// TIA Portal project "DHARMA_1500" (V15) (continued)
VAR_GLOBAL   // PLC tag table "VAT_DeSelectModule"
   "HM_DP_Bus_MK01_Melden" AT %M30.0 : Bool;
   "HM_DP_Bus_MK01_speichern" AT %M30.1 : Bool;
   "HM_DP_Bus_MK01_aktiv" AT %M30.2 : Bool;
   "HM_DP_Bus_MK02_Melden" AT %M30.3 : Bool;
   "HM_DP_Bus_MK02_speichern" AT %M30.4 : Bool;
   "HM_DP_Bus_MK02_aktiv" AT %M30.5 : Bool;
   "HM_DP_Bus_MK03_Melden" AT %M30.6 : Bool;
   "HM_DP_Bus_MK03_speichern" AT %M30.7 : Bool;
   "HM_DP_Bus_MK03_aktiv" AT %M31.0 : Bool;
   "HM_DP_Bus_MK04_Melden" AT %M31.1 : Bool;
   "HM_DP_Bus_MK04_speichern" AT %M31.2 : Bool;
   "HM_DP_Bus_MK04_aktiv" AT %M31.3 : Bool;
   "HM_DP_Bus_MK05_Melden" AT %M31.4 : Bool;
   "HM_DP_Bus_MK05_speichern" AT %M31.5 : Bool;
   "HM_DP_Bus_MK05_aktiv" AT %M31.6 : Bool;
   "HM_DP_Bus_MK06_Melden" AT %M31.7 : Bool;
   "HM_DP_Bus_MK06_speichern" AT %M32.0 : Bool;
   "HM_DP_Bus_MK06_aktiv" AT %M32.1 : Bool;
   "HM_DP_Bus_MK07_Melden" AT %M32.2 : Bool;
   "HM_DP_Bus_MK07_speichern" AT %M32.3 : Bool;
   "HM_DP_Bus_MK07_aktiv" AT %M32.4 : Bool;
   "HM_DP_Bus_MK08_Melden" AT %M32.5 : Bool;
   "HM_DP_Bus_MK08_speichern" AT %M32.6 : Bool;
   "HM_DP_Bus_MK08_aktiv" AT %M32.7 : Bool;
   "HM_DP_Bus_MK09_Melden" AT %M33.0 : Bool;
   "HM_DP_Bus_MK09_speichern" AT %M33.1 : Bool;
   "HM_DP_Bus_MK09_aktiv" AT %M33.2 : Bool;
   "HM_DP_Bus_MK10_Melden" AT %M33.3 : Bool;
   "HM_DP_Bus_MK10_speichern" AT %M33.4 : Bool;
   "HM_DP_Bus_MK10_aktiv" AT %M33.5 : Bool;
   "HM_DP_Bus_MK11_Melden" AT %M33.6 : Bool;
   "HM_DP_Bus_MK11_speichern" AT %M33.7 : Bool;
   "HM_DP_Bus_MK11_aktiv" AT %M34.0 : Bool;
   "HM_DP_Bus_MK12_Melden" AT %M34.1 : Bool;
   "HM_DP_Bus_MK12_speichern" AT %M34.2 : Bool;
   "HM_DP_Bus_MK12_aktiv" AT %M34.3 : Bool;
   "HM_DP_Bus_MK13_Melden" AT %M34.4 : Bool;
   "HM_DP_Bus_MK13_speichern" AT %M34.5 : Bool;
   "HM_DP_Bus_MK13_aktiv" AT %M34.6 : Bool;
   "HM_DP_Bus_MK14_Melden" AT %M34.7 : Bool;
   "HM_DP_Bus_MK14_speichern" AT %M35.0 : Bool;
   "HM_DP_Bus_MK14_aktiv" AT %M35.1 : Bool;
   "HM_DP_Bus_MK15_Melden" AT %M35.2 : Bool;
   "HM_DP_Bus_MK15_speichern" AT %M35.3 : Bool;
   "HM_DP_Bus_MK15_aktiv" AT %M35.4 : Bool;
   "HM_DP_An_Abmelden_Busy" AT %M29.7 : Bool;
END_VAR

VAR_GLOBAL   // PLC tag table "Robots"
   "FHM_PU_cycle_running" AT %M850.0 : Bool;
   "Flag_PU_cycle_running" AT %M850.1 : Bool;
END_VAR

VAR_GLOBAL   // PLC tag table "VAT_VB_Skripte"
   "new_shift" AT %M4.0 : Bool;
   "flag_delay_check_path" AT %M7.1 : Bool;
   "Flag_Network" AT %M1.7 : Bool;
END_VAR

VAR_GLOBAL   // PLC tag table "Shot_protocol"
   "M_ShotActive" AT %M1002.3 : Bool;
   "TotalFlowShotC01" AT %MD950 : Real;
   "TotalFlowShotC02" AT %MD954 : Real;
   "TotalFlowShotC03" AT %MD958 : Real;
   "TotalFlowShotC04" AT %MD962 : Real;
   "TotalFlowShotC05" AT %MD966 : DInt;
   "TotalFlowShotC06" AT %MD970 : DInt;
   "TotalFlowShotC07" AT %MD974 : DInt;
   "TotalFlowShotC08" AT %MD978 : DInt;
   "TotalFlowShotC09" AT %MD982 : DInt;
   "TotalFlowShotC10" AT %MD986 : DInt;
   "TotalFlowShotC11" AT %MD990 : DInt;
   "TotalFlowShotC12" AT %MD994 : DInt;
   "CompAtShot" AT %MW942 : Word;
   "AmountFlowValuesMa1C1" AT %MD800 : Real;
   "AmountFlowValuesMa1C2" AT %MD804 : Real;
   "AmountFlowValuesMa1C3" AT %MD808 : Real;
   "AmountFlowValuesMa1C4" AT %MD812 : Real;
   "FHF_ShotreleaseM1" AT %M940.2 : Bool;
   "M1C01active" AT %M932.0 : Bool;
   "M1C02active" AT %M932.1 : Bool;
   "M1C03active" AT %M932.2 : Bool;
   "M1C04active" AT %M932.3 : Bool;
   "HF_FP_ShotRuns" AT %M941.0 : Bool;
   "HF_FP_ShotStoppedM1" AT %M940.4 : Bool;
   "BufferShotResultM1" AT %M920.0 : Bool;
   "FHM_ShotRunsMH1" AT %M402.0 : Bool;
   "FP_BufferShotResultM1" AT %M919.0 : Bool;
   "M1C05active" AT %M932.4 : Bool;
   "M1C06active" AT %M932.5 : Bool;
   "M1C07active" AT %M932.6 : Bool;
   "M1C08active" AT %M932.7 : Bool;
   "M1C09active" AT %M933.0 : Bool;
   "M1C10active" AT %M933.1 : Bool;
   "M1C11active" AT %M933.2 : Bool;
   "M1C12active" AT %M933.3 : Bool;
   "AmountFlowValuesMa1C5" AT %MD816 : Real;
   "AmountFlowValuesMa1C6" AT %MD820 : Real;
   "AmountFlowValuesMa1C7" AT %MD824 : Real;
   "AmountFlowValuesMa1C8" AT %MD828 : Real;
   "AmountFlowValuesMa1C9" AT %MD832 : Real;
   "AmountFlowValuesMa1C10" AT %MD836 : Real;
   "AmountFlowValuesMa1C11" AT %MD840 : Real;
   "AmountFlowValuesMa1C12" AT %MD844 : Real;
END_VAR

VAR_GLOBAL   // PLC tag table "All_other"
   "TT_Quitt_Door_1" AT %I1102.1 : Bool;
   "TT_H_Empty" AT %Q104.5 : Bool;
   "TT_H_WithoutFoam" AT %Q104.6 : Bool;
   "K_TraceHeatingM1C4" AT %Q16.6 : Bool;
   "Flag_Req_read_DPBus_01" AT %M9.0 : Bool;
   "Flag_Req_read_DP1_Busy" AT %M9.1 : Bool;
   "Flag_Req_read_IO_Busy" AT %M9.2 : Bool;
   "HF_FLT_QPB_C1" AT %M120.1 : Bool;
   "HF_FLT_QPB_C2" AT %M120.2 : Bool;
   "HF_FLT_QPB_C3" AT %M120.3 : Bool;
   "HF_FLT_QPB_C4" AT %M120.4 : Bool;
   "F_CycleRunningMH01" AT %M390.0 : Bool;
   "F_CycleRunningMH02" AT %M390.1 : Bool;
   "F_CycleRunningMH03" AT %M390.2 : Bool;
   "F_CycleRunningMH04" AT %M390.3 : Bool;
   "F_CycleRunningMH05" AT %M390.4 : Bool;
   "F_CycleRunningMH06" AT %M390.5 : Bool;
   "F_CycleRunningMH07" AT %M390.6 : Bool;
   "F_CycleRunningMH08" AT %M390.7 : Bool;
   "StopShotCorrMH01" AT %M309.4 : Bool;
   "StopShotCorrMH02" AT %M309.5 : Bool;
   "StopShotCorrMH03" AT %M309.6 : Bool;
   "StopShotCorrMH04" AT %M309.7 : Bool;
   "ShotFinishedModul_MH01" AT %M122.1 : Bool;
   "ShotFinishedModul_MH02" AT %M122.2 : Bool;
   "ShotFinishedModul_MH03" AT %M122.3 : Bool;
   "ShotFinishedModul_MH04" AT %M122.4 : Bool;
   "ShotFinishedModul_MH05" AT %M122.5 : Bool;
   "ShotFinishedModul_MH06" AT %M122.6 : Bool;
   "ShotFinishedModul_MH07" AT %M122.7 : Bool;
   "ShotFinishedModul_MH08" AT %M123.0 : Bool;
   "ShotFinishedModul_MH09" AT %M123.1 : Bool;
   "ShotFinishedModul_MH10" AT %M123.2 : Bool;
   "ShotFinishedModul_MH11" AT %M123.3 : Bool;
   "ShotFinishedModul_MH12" AT %M123.4 : Bool;
   "ShotFinishedModul_MH13" AT %M123.5 : Bool;
   "ShotFinishedModul_MH14" AT %M123.6 : Bool;
   "ShotFinishedModul_MH15" AT %M123.7 : Bool;
   "ShotFinishedModul_MH16" AT %M124.0 : Bool;
   "EnableFinishShot_MH01" AT %M106.0 : Bool;
   "EnableFinishShot_MH02" AT %M106.1 : Bool;
   "EnableFinishShot_MH03" AT %M106.2 : Bool;
   "EnableFinishShot_MH04" AT %M106.3 : Bool;
   "EnableFinishShot_MH05" AT %M106.4 : Bool;
   "EnableFinishShot_MH06" AT %M106.5 : Bool;
   "EnableFinishShot_MH07" AT %M106.6 : Bool;
   "EnableFinishShot_MH08" AT %M106.7 : Bool;
   "ShotNoNextMa1" AT %MW556 : Int;
   "ShotNoNextMa2" AT %MW558 : Int;
   "ShotNoNextMa3" AT %MW560 : Int;
   "ShotNoNextMa4" AT %MW562 : Int;
   "StopShotCorrMH08" AT %M319.7 : Bool;
   "StopShotCorrMH07" AT %M319.6 : Bool;
   "StopShotCorrMH06" AT %M319.5 : Bool;
   "StopShotCorrMH05" AT %M319.4 : Bool;
   "CalcShotValuesMa1" AT %M135.0 : Bool;
   "ShotStoppedM1" AT %M135.1 : Bool;
   "M1200_ActivateAdrProCan" AT %M120.0 : Bool;
   "NoShotActiveM1" AT %M158.0 : Bool;
   "F_CycleRunningMH09" AT %M391.0 : Bool;
   "F_CycleRunningMH10" AT %M391.1 : Bool;
   "F_CycleRunningMH11" AT %M391.2 : Bool;
   "F_CycleRunningMH12" AT %M391.3 : Bool;
   "F_CycleRunningMH13" AT %M391.4 : Bool;
   "F_CycleRunningMH14" AT %M391.5 : Bool;
   "F_CycleRunningMH15" AT %M391.6 : Bool;
   "F_CycleRunningMH16" AT %M391.7 : Bool;
   "StopShotCorrMH10" AT %M320.1 : Bool;
   "StopShotCorrMH09" AT %M320.0 : Bool;
   "Start_Controler1_HP_K1" AT %M180.5 : Bool;
   "Start_Controler2_HP_K1" AT %M180.4 : Bool;
   "Start_Controler1_HP_K2" AT %M181.5 : Bool;
   "Start_Controler2_HP_K2" AT %M181.4 : Bool;
   "Start_Controler2_LP_K1" AT %M182.4 : Bool;
   "Start_Controler1_LP_K1" AT %M182.5 : Bool;
   "Start_Controler2_LP_K2" AT %M183.4 : Bool;
   "Start_Controler1_LP_K2" AT %M183.5 : Bool;
   "Flag_ToggleForDatarequest" AT %M2.7 : Bool;
   "FP_new_page_no" AT %M566.0 : Bool;
   "PulsShotend_M1_MH_No" AT %MW201 : Word;
   "NextShot_M1_MH_No" AT %MW212 : Word;
   "HM_FP_ShotFound_M1" AT %M370.0 : Bool;
END_VAR

VAR_GLOBAL   // PLC tag table "Timer"
   "TM_WatchdogProcan01" AT %T150 : Timer;
   "TM_WatchdogProcan02" AT %T151 : Timer;
   "TM_WatchdogProcan03" AT %T152 : Timer;
   "TM_WatchdogProcan04" AT %T153 : Timer;
   "TM_WatchdogProcan05" AT %T154 : Timer;
   "TM_WatchdogProcan06" AT %T155 : Timer;
   "TM_WatchdogProcan07" AT %T156 : Timer;
   "TM_WatchdogProcan08" AT %T157 : Timer;
   "TM_WatchdogProcan09" AT %T158 : Timer;
   "TM_WatchdogProcan10" AT %T159 : Timer;
   "TM_WatchdogProcan11" AT %T149 : Timer;
   "TM_HP_after_shot_M1" AT %T12 : Timer;
   "TM_Kreislauf_ND_M1" AT %T42 : Timer;
   "TM_OM_M1" AT %T10 : Timer;
   "TM_Kreislauf_M1" AT %T11 : Timer;
   "TM_P_oben_MK_Hyd_M1" AT %T20 : Timer;
   "TM_MK_Hyd_Temp_M1" AT %T22 : Timer;
   "TM_MK_Hyd_M1" AT %T24 : Timer;
   "TM_MK_Hyd_Filter_M1" AT %T23 : Timer;
   "TM_SwitchOffHydMH_M1" AT %T21 : Timer;
   "TM_USE_Taktzeit_M1" AT %T40 : Timer;
   "TM_USE_Umschaltzeit_M1" AT %T41 : Timer;
   "TM_SwitchOnDelayFCPump" AT %T26 : Timer;
   "TM_EdgeFilter01" AT %T54 : Timer;
   "TM1_FeedPump01" AT %T55 : Timer;
   "TM2_FeedPump01" AT %T60 : Timer;
   "TM_RestartC01" AT %T56 : Timer;
   "TM_CtrlFeedPumpC01" AT %T57 : Timer;
   "TM_CommonC01" AT %T58 : Timer;
   "TM_DelayClosedLoopC01" AT %T59 : Timer;
   "TM_IntervalC01" AT %T61 : Timer;
   "TM_EdgeFilter02" AT %T62 : Timer;
   "TM1_FeedPump02" AT %T63 : Timer;
   "TM_RestartC02" AT %T64 : Timer;
   "TM_CtrlFeedPumpC02" AT %T65 : Timer;
   "TM_CommonC02" AT %T66 : Timer;
   "TM_DelayClosedLoopC02" AT %T67 : Timer;
   "TM2_FeedPump02" AT %T68 : Timer;
   "TM_IntervalC02" AT %T69 : Timer;
   "TM_RunTime_CP01" AT %T30 : Timer;
   "TM_RunTime_CP02" AT %T31 : Timer;
   "TM_RunTime_CP03" AT %T32 : Timer;
   "TM_RunTime_CP04" AT %T33 : Timer;
   "TM_RunTime_CP05" AT %T34 : Timer;
   "TM_RunTime_CP06" AT %T35 : Timer;
   "TM_RunTime_CP07" AT %T36 : Timer;
   "TM_RunTime_CP08" AT %T37 : Timer;
   "TM_FltCPHomePos_CP01" AT %T241 : Timer;
   "TM_FltCPHomePos_CP02" AT %T242 : Timer;
   "TM_FltCPHomePos_CP03" AT %T243 : Timer;
   "TM_FltCPHomePos_CP04" AT %T244 : Timer;
   "TM_FltCPHomePos_CP05" AT %T245 : Timer;
   "TM_FltCPHomePos_CP06" AT %T246 : Timer;
   "TM_FltCPHomePos_CP07" AT %T247 : Timer;
   "TM_FltCPHomePos_CP08" AT %T248 : Timer;
   "TM_HydrForCPoffM1" AT %T226 : Timer;
   "TM_CycleTimer_M1" AT %T39 : Timer;
   "TM_Vac1DelayLock" AT %T100 : Timer;
   "TM_Vac2DelayLock" AT %T101 : Timer;
   "TM_Vac1DelayPump" AT %T102 : Timer;
   "TM_Vac2DelayPump" AT %T103 : Timer;
   "TM1_Agitator_01" AT %T160 : Timer;
   "TM2_Agitator_01" AT %T161 : Timer;
   "TM1_Agitator_02" AT %T162 : Timer;
   "TM2_Agitator_02" AT %T163 : Timer;
   "TM_Refilling_01" AT %T168 : Timer;
   "TM_Refilling_02" AT %T169 : Timer;
   "TM1_Agitator_03" AT %T164 : Timer;
   "TM2_Agitator_03" AT %T165 : Timer;
   "TM_Refilling_03" AT %T170 : Timer;
   "TM1_Charge_C3" AT %T166 : Timer;
   "TM2_Charge_C3" AT %T167 : Timer;
   "TM_FltCPHomePos_CP09" AT %T249 : Timer;
   "TM_FltCPHomePos_CP10" AT %T250 : Timer;
   "TM_RunTime_CP09" AT %T38 : Timer;
   "TM_RunTime_CP10" AT %T43 : Timer;
   "TM_FanPumpC01" AT %T220 : Timer;
   "TM_delay_2PointAdjust_C1" AT %T70 : Timer;
   "TM_delay_2PointAdjust_C2" AT %T71 : Timer;
   "TM_Interrupt2PointAdjustment" AT %T27 : Timer;
   "TM_pulse_2PointAdjust_C1" AT %T28 : Timer;
   "TM_pulse_2PointAdjust_C2" AT %T29 : Timer;
   "T_Delay_Send_Data_KMI" AT %T251 : Timer;
   "TIM_Spuelzeit" AT %T216 : Timer;
   "TIM_Delay_flushing" AT %T217 : Timer;
   "TM_Max_Wartezeit_MKR2" AT %T215 : Timer;
   "TM_Delay_Cleaning_man" AT %T218 : Timer;
   "TIM_Delay_Clean_air" AT %T219 : Timer;
   "TIM_Delay_Blow_Air" AT %T224 : Timer;
   "TM_1_Robot_1" AT %T230 : Timer;
   "TM_2_Robot_1" AT %T231 : Timer;
   "TM_3_Robot_1" AT %T232 : Timer;
   "TM_4_Robot_1" AT %T233 : Timer;
   "TM_5_Robot_1" AT %T234 : Timer;
   "TM_6_Robot_1" AT %T235 : Timer;
   "TM_7_Robot_1" AT %T236 : Timer;
   "TMTT_OPMode" AT %T1406 : Timer;
   "TMTT_StartProduction" AT %T1407 : Timer;
   "TMTT_Production" AT %T1408 : Timer;
   "TMTT_Tact" AT %T1409 : Timer;
   "TMTT_IPOS_Universal" AT %T1410 : Timer;
   "TMTT_IPOS_Enable" AT %T1411 : Timer;
   "TMTT_IPOS_TolInPos" AT %T1412 : Timer;
   "TMTT_IPOS_FaultFC" AT %T1413 : Timer;
   "TMTT_IPOS_DelayInPos" AT %T1414 : Timer;
   "TMTT_IPOS_Horn" AT %T1415 : Timer;
   "TMTT_RunTimeManipulator" AT %T1416 : Timer;
   "TMTT_WaitTimeMHFront" AT %T1417 : Timer;
   "TMTT_RunTimeCPCleaner" AT %T1418 : Timer;
   "TMTT_DelayMHCleaning" AT %T1419 : Timer;
   "TMTT_DuringMHCleaning" AT %T1420 : Timer;
   "delay_timer" AT %T4 : Timer;
   "Timer_Network" AT %T5 : Timer;
   "Timer_Network_reset" AT %T6 : Timer;
   "Timer_check_path" AT %T7 : Timer;
   "TM_DelayEmergencyStop" AT %T228 : Timer;
   "TM_Tank_Delay_DryRun_FeedPump_C1" AT %T200 : Timer;
   "TM_Tank_Delay_DryRun_FeedPump_C2" AT %T201 : Timer;
   "TM_ExhauseSystem" AT %T210 : Timer;
   "TM_Overlap_Valves_Pentan" AT %T211 : Timer;
   "TM_Valve1_Pentan" AT %T212 : Timer;
   "TM_Valve2_Pentan" AT %T213 : Timer;
   "T_Leakage_Ctrl_N2" AT %T180 : Timer;
   "T_Leakage_Ctrl_Tact_N2" AT %T181 : Timer;
   "T_Inerting" AT %T182 : Timer;
   "T_Ready_for_Shot" AT %T183 : Timer;
   "T_Delay_Purge" AT %T184 : Timer;
   "T_Purge" AT %T185 : Timer;
   "T_Max_Inerting" AT %T186 : Timer;
   "T_Delay_Plunger" AT %T187 : Timer;
   "T_Delay_Purge_Tact" AT %T188 : Timer;
   "T_Purge_Tact" AT %T189 : Timer;
   "T_Pause_Tact" AT %T190 : Timer;
   "T_Total_Time_Purge" AT %T191 : Timer;
   "TM_Reset_after_purge" AT %T194 : Timer;
   "TM_Purge_after_Shot" AT %T195 : Timer;
   "TM_Nozzle_off_delay_MH01" AT %T252 : Timer;
   "TM_FanPumpC02" AT %T221 : Timer;
   "TM_Delay_nozzle_off_MH1" AT %T253 : Timer;
   "TM_RFID_ready_MH1" AT %T132 : Timer;
   "TM_RFID_ready_MH2" AT %T133 : Timer;
   "TM_Verz_Sync_1" AT %T199 : Timer;
   "TM_Delay_Limit_Control" AT %T2 : Timer;   // At the opening from the mixinghead wait with checking the limits
   "TM_Alarm_QPBTime_C1" AT %T1 : Timer;
   "TM_Alarm_QPBTime_C2" AT %T3 : Timer;
   "TM_Betriebsart_Anlage" AT %T1421 : Timer;
   "TM_Anfahrwarnung_Anlage" AT %T1422 : Timer;
   "TM_Produktion_Anlage" AT %T1423 : Timer;
   "TM_Ansteuerung_SEW" AT %T1424 : Timer;
   "TM_Nachlauf_Freigabe_SEW" AT %T1425 : Timer;
   "TM_Verz_STG_Genauhalt" AT %T1426 : Timer;
   "TM_Delay_target_reached" AT %T1427 : Timer;
   "TM_Delay_autostop_okay_FC" AT %T1428 : Timer;
   "TM_SV_Quitt_Fault" AT %T1429 : Timer;
   "TM_STG_Kettenentlastung" AT %T1430 : Timer;
   "TM_Kettenspanner" AT %T1431 : Timer;
   "TM_Taktzeit" AT %T1432 : Timer;
   "TM_CS_K2" AT %T80 : Timer;
   "TIM_FRA_WDG1" AT %T8 : Timer;
   "TIM_FRA_WDG2" AT %T9 : Timer;
   "TM_Delay_Safetydoor_1" AT %T237 : Timer;
   "TM_Delay_Safetydoor_2" AT %T238 : Timer;
   "TM_Hydraulik_RK_Druck" AT %T13 : Timer;
   "T_Set_new_page_no" AT %T14 : Timer;
   "TM_Group1_Fault" AT %T500 : Timer;
END_VAR

VAR_GLOBAL   // PLC tag table "Counter"
   "Z_HubzaehlerM1" AT %C10 : Counter;
   "CT_MK_Reinigungen_MK2" AT %C15 : Counter;
END_VAR

VAR_GLOBAL   // PLC tag table "VAT_Trace"
   "M_NewShotDataToMC" AT %M587.6 : Bool;
   "M_NewShotDataToMC_01" AT %M700.1 : Bool;
   "M_WriteShotDataMC_01" AT %M704.0 : Bool;
   "M_FP_NewShotDataToMC_01" AT %M700.0 : Bool;
   "M_FP_NewShotDataToMC_02" AT %M700.2 : Bool;
   "M_NewShotDataToMC_02" AT %M700.3 : Bool;
   "M_WriteShotDataMC_02" AT %M704.1 : Bool;
   "HF_new_shot_data" AT %M587.7 : Bool;
   "HT_new_shot_data_valid" AT %M588.0 : Bool;
   "M_WriteShotDataMC_03" AT %M704.2 : Bool;
   "M_WriteShotDataMC_04" AT %M704.3 : Bool;
   "M_WriteShotDataTestShot" AT %M704.4 : Bool;
   "M_FP_NewShotDataToMC_03" AT %M700.4 : Bool;
   "M_NewShotDataToMC_03" AT %M700.5 : Bool;
   "M_FP_NewShotDataToMC_04" AT %M700.6 : Bool;
   "M_NewShotDataToMC_04" AT %M700.7 : Bool;
   "M_FP_NewShotDataTestShot" AT %M701.0 : Bool;
   "M_NewShotDataTestShot" AT %M701.1 : Bool;
   "TM_FLT_Com_DataShot_MC01" AT %T432 : Timer;
   "TM_FLT_Com_DataShot_MC02" AT %T433 : Timer;
   "TM_FLT_Com_DataShot_MC03" AT %T434 : Timer;
   "TM_FLT_Com_DataShot_MC04" AT %T435 : Timer;
END_VAR

TYPE "UDT1004_MH_Status"
VERSION : 0.1
   STRUCT
      SWU_released : Bool;
      SWU_activ : Bool;
      QPB_Values_selected : Bool;
      LP_Exist : Bool;
      Indicator_HP : Bool;
      Switch_HP_ON_OFF : Bool;
      Switch_Service_ON_OFF : Bool;
      FaultExist : Bool;
      OpenMHEnableExtern : Bool;   // External enable to open the mixinghead
      Switch_Testshot_A_ON_OFF : Bool;
      Switch_Testshot_B_ON_OFF : Bool;
      Spare11 : Bool;
      Spare12 : Bool;
      Spare13 : Bool;
      Spare14 : Bool;
      Spare15 : Bool;
      State_HP : Int;
      State_Service : Int;
      State_Testshot_A : Int;
      State_Testshot_B : Int;
   END_STRUCT;
END_TYPE

TYPE "UDT002_Word_1_16"
VERSION : 0.0
   STRUCT
      "09" : Bool;   // ... Nummer 09 ist angewählt/ aktiv etc.
      "10" : Bool;   // ... Nummer 10 ist angewählt/ aktiv etc.
      "11" : Bool;   // ... Nummer 11 ist angewählt/ aktiv etc.
      "12" : Bool;   // ... Nummer 12 ist angewählt/ aktiv etc.
      "13" : Bool;   // ... Nummer 13 ist angewählt/ aktiv etc.
      "14" : Bool;   // ... Nummer 14 ist angewählt/ aktiv etc.
      "15" : Bool;   // ... Nummer 15 ist angewählt/ aktiv etc.
      "16" : Bool;   // ... Nummer 16 ist angewählt/ aktiv etc.
      "01" : Bool;   // ... Nummer 01 ist angewählt/ aktiv etc.
      "02" : Bool;   // ... Nummer 02 ist angewählt/ aktiv etc.
      "03" : Bool;   // ... Nummer 03 ist angewählt/ aktiv etc.
      "04" : Bool;   // ... Nummer 04 ist angewählt/ aktiv etc.
      "05" : Bool;   // ... Nummer 05 ist angewählt/ aktiv etc.
      "06" : Bool;   // ... Nummer 06 ist angewählt/ aktiv etc.
      "07" : Bool;   // ... Nummer 07 ist angewählt/ aktiv etc.
      "08" : Bool;   // ... Nummer 08 ist angewählt/ aktiv etc.
   END_STRUCT;
END_TYPE

TYPE "UDT001_DWord_1_32"
VERSION : 0.0
   STRUCT
      "25" : Bool;   // ... Number 25 is selected and active
      "26" : Bool;   // ... Number 26 is selected and active
      "27" : Bool;   // ... Number 27 is selected and active
      "28" : Bool;   // ... Number 28 is selected and active
      "29" : Bool;   // ... Number 29 is selected and active
      "30" : Bool;   // ... Number 30 is selected and active
      "31" : Bool;   // ... Number 31 is selected and active
      "32" : Bool;   // ... Number 32 is selected and active
      "17" : Bool;   // ... Number 17 is selected and active
      "18" : Bool;   // ... Number 18 is selected and active
      "19" : Bool;   // ... Number 19 is selected and active
      "20" : Bool;   // ... Number 20 is selected and active
      "21" : Bool;   // ... Number 21 is selected and active
      "22" : Bool;   // ... Number 22 is selected and active
      "23" : Bool;   // ... Number 23 is selected and active
      "24" : Bool;   // ... Number 24 is selected and active
      "09" : Bool;   // ... Number 09 is selected and active
      "10" : Bool;   // ... Number 10 is selected and active
      "11" : Bool;   // ... Number 11 is selected and active
      "12" : Bool;   // ... Number 12 is selected and active
      "13" : Bool;   // ... Number 13 is selected and active
      "14" : Bool;   // ... Number 14 is selected and active
      "15" : Bool;   // ... Number 15 is selected and active
      "16" : Bool;   // ... Number 16 is selected and active
      "01" : Bool;   // ... Number 01 is selected and active
      "02" : Bool;   // ... Number 02 is selected and active
      "03" : Bool;   // ... Number 03 is selected and active
      "04" : Bool;   // ... Number 04 is selected and active
      "05" : Bool;   // ... Number 05 is selected and active
      "06" : Bool;   // ... Number 06 is selected and active
      "07" : Bool;   // ... Number 07 is selected and active
      "08" : Bool;   // ... Number 08 is selected and active
   END_STRUCT;
END_TYPE

TYPE "UDT925_Shot"
VERSION : 0.1
   STRUCT
      MHNo : Int := 0;   // Mixinghead number
      FoamingTime : Real := 100.0;   // Foaming Time
      PartWeight : Real := 200.0;   // Part Weight
      CP_ThrottleGap : Real;   // Throttle gap of an analog cleaning piston
      SwitchOff_Pressure : Real;   // Pressure to switch off foaming cycle
      PartCounter : Int;   // Number of PartCounter
      Pressure : Array[1..6] of Real;   // Pressure for 6 components
      Flow : Array[1..6] of Real;   // Flow for 6 components
      RefComponent : Int;   // Number of the reference component
      PartShotDisable : Bool;   // Disable foaming
      CPMoveAfterShot : Bool;   // Cleaning piston moves after shot
      PurgeMHAfterShot : Bool;   // Cleaning mixhead direct after shot with air or nitrogen
      "2PoinMovement_Comp01" : Bool;
      "2PoinMovement_Comp02" : Bool;
      "2PoinMovement_Comp03" : Bool;
      "2PoinMovement_Comp04" : Bool;
      "2PoinMovement_Comp05" : Bool;
      "2PoinMovement_Comp06" : Bool;
      Spare_1 : Bool;
      Spare_2 : Bool;
      Spare_3 : Bool;
      Spare_4 : Bool;
      Spare_5 : Bool;
      Spare_6 : Bool;
      Spare_7 : Bool;
   END_STRUCT;
END_TYPE

TYPE "UDT885_AnaChannel"
VERSION : 0.1
   STRUCT
      Channal : Array[1..8] of "UDT901_ConfAna";
   END_STRUCT;
END_TYPE

TYPE "UDT930_Tool"
TITLE = Foaming: Tool set values RAM
VERSION : 0.1
   STRUCT
      tool_name : String[20];   // name of tool
      Rob_Prog : Int;   // Robot program number 1
      Rob_Prog2 : Int;   // Robot program number 2
      PartShot_Amount : Byte := B#16#0;   // Amount of part shoots at this tool
      RefComponent : Byte;   // Number of the reference component
      Spare : Byte;
      EnableTool : Bool;   // Enable Bit: tool should be foamed
      Spare5_2 : Bool;
      Spare5_3 : Bool;
      Spare5_4 : Bool;
      Spare5_5 : Bool;
      Spare5_6 : Bool;
      EnablePurgeMH : Bool;   // Enable Bit: Mixhead cleaning with air or nitrogen
      NitrogenVol : Int;   // Nitrogen volume complete
      Spare_12 : Word := W#16#0;
   END_STRUCT;
END_TYPE

TYPE "UDT932_SaveProg"
VERSION : 0.1
   STRUCT
      ProgramNo : Int;
   END_STRUCT;
END_TYPE

TYPE "UDT926_ShotSet"
VERSION : 0.1
   STRUCT
      Shot : Array[1.."AmountPartShots"] of "UDT925_Shot";
   END_STRUCT;
END_TYPE

TYPE "UDT937_ShotData"
VERSION : 0.1
   STRUCT
      MH_Conn_at_shot : Byte;   // MH connections which are involved at this shot (Bit 0 - 7 -> Connection 1 - 8)
      MH_No : Byte;   // Mixinghead no. at shot
      Comp_at_Shot : Word;   // Component which are involved at this shot (Bit 0-11 -> Comp 1-12)
      PartCounter : Int;   // Actual Part counter // per mould or per PartShot
      CP_AfterShot : Bool;   // Cleaning stroke after shot selected
      PurgeMH_AfterShot : Bool;   // Cleaning MH with air or nitrogen after shot
      ShotDisabled : Bool;   // The selected shot is disabled -> like service shot
      Spare03 : Bool;
      Spare04 : Bool;
      Spare05 : Bool;
      Spare06 : Bool;
      Spare07 : Bool;
      Spare08 : Bool;
      Spare09 : Bool;
      Spare10 : Bool;
      Spare11 : Bool;
      Spare12 : Bool;
      Spare13 : Bool;
      Spare14 : Bool;
      Spare15 : Bool;
      Foamingtime : Real;
      Flow : Array[1..6] of Real;   // Flowrates of the material (1/100 g/s) at mixinghead connection (1-6)
      Pressure : Array[1..6] of Real;   // Setvalues of pressure of material at mixinghead connection (1-6)
      "2PointAdjustment" : Array[1..8] of Bool;   // Selection for 2- Point Adjustment at mixinghead connection (1-6)
   END_STRUCT;
END_TYPE

TYPE "UDT10_Machine"
TITLE = State of machine please customize
VERSION : 0.1
   STRUCT
      HydStartUp_finished : Bool;   // All at the machine used hydraulic units are running and OK
      HP_after_shot : Bool;   // Activate highpressure circualtion after a automatic shot
      Flag_P_HP_after_shot : Bool;   // Flag switch on high pressure circulation after shot
      Flag_N_HP_after_shot : Bool;   // Flag switch off high pressure circulation after shot
      Flag_N_HP_partner : Bool;   // Flankenmerker zum löschen der Pausenzeit bei der Partneranlage
      Reserve_0_5 : Bool;
      Reserve_0_6 : Bool;
      Reserve_0_7 : Bool;
      Fault_Cooling_MH_Hydr : Bool;   // Fault: cooling mixinghead hydraulic
      Fault_filter_Cooling_Hyd : Bool;   // Fault: Back flow filter cooling mixinghead hydraulic
      Fault_P_max_Hydr : Bool;   // Fault: Max. pressure edge filter mixinghead hydraulic
      Reserve_1_3 : Bool;
      Fault_Fillingpump_K1 : Bool;   // Fault: Filling pump daytank Poly 1
      Fault_Fillingpump_K2 : Bool;   // Fault: Filling pump daytank Iso
      Fault_Fillingpump_K3 : Bool;   // Fault: Filling pump daytank Poly 2
      Fault_Fillingpump_K4 : Bool;   // Fault: Filling pump daytank Poly 3
      Metering : "UDT002_Word_1_16";   // Komponenten- Nummer die dosiert werden soll
   END_STRUCT;
END_TYPE

TYPE "UDT011_Operationmode"
TITLE = State of operation mode machine
VERSION : 0.0
   STRUCT
      valid : Bool;   // A valid operation mode is selected (manual or automatic)
      Manual : Bool;   // Control voltage on and manual mode selected
      Auto : Bool;   // Control voltage on and automatic mode selected
      Cylinderservice : Bool;   // Cylinder service and manual mode selected and no recirculation active
      Test : Bool;   // Operation mode automatic and test selected // Test pouring by test valves
      Operation : Bool;   // Operation mode without foam (Service) to test the pouring sequence
      Lamptest : Bool;   // Controlvoltage on and lamp test active
      Controllvoltage : Bool;   // Signal "Controlvoltage ON" is more than 1s active
      Edge_OM_Change : Bool;   // Edge flag switch over between service/operation mode
      Active : Bool;   // A valid operation mode was selected and hydraulic is active
      SwitchManual : Bool;   // Switch manual from external plant
      SwitchAutomatic : Bool;   // Switch automatic from external plant
      SwitchOperation : Bool;   // Switch operation mode ->ON -> with foam to open mixinghead (extarnel)
      SwitchWeekEnd : Bool;   // Switch WeekEnd Mode is selected
      SwitchLamptest : Bool;   // Switch Lamptest is selected
      Spare16 : Bool;
   END_STRUCT;
END_TYPE

